// TIA Portal project "Linie_reciclare_paleti_mod" (V16) (continued)
               Length : Int := 1;
               BlockStat : DWord;
               IOLStat : DWord;
               RelRead : Bool := TRUE;
               RelWrite : Bool := TRUE;
            END_STRUCT;
            Parameter_13 : Struct
               V_X1_3_DO2Sub8 : Byte := BYTE#16#00;
               Byte01 : Byte := BYTE#16#00;
               Byte02 : Byte := BYTE#16#00;
               Byte03 : Byte := BYTE#16#00;
               Index : Int := 15000;
               Subindex : Int := 8;
               Length : Int := 1;
               BlockStat : DWord;
               IOLStat : DWord;
               RelRead : Bool := TRUE;
               RelWrite : Bool := TRUE;
            END_STRUCT;
            Parameter_14 : Struct
               V_X1_4_DO1Sub9 : Byte := BYTE#16#00;
               Byte01 : Byte := BYTE#16#00;
               Byte02 : Byte := BYTE#16#00;
               Byte03 : Byte := BYTE#16#00;
               Index : Int := 15000;
               Subindex : Int := 9;
               Length : Int := 1;
               BlockStat : DWord;
               IOLStat : DWord;
               RelRead : Bool := TRUE;
               RelWrite : Bool := TRUE;
            END_STRUCT;
            Parameter_15 : Struct
               V_X1_4_DO2Sub10 : Byte := BYTE#16#00;
               Byte01 : Byte := BYTE#16#00;
               Byte02 : Byte := BYTE#16#00;
               Byte03 : Byte := BYTE#16#00;
               Index : Int := 15000;
               Subindex : Int := 10;
               Length : Int := 1;
               BlockStat : DWord;
               IOLStat : DWord;
               RelRead : Bool := TRUE;
               RelWrite : Bool := TRUE;
            END_STRUCT;
            Parameter_16 : Struct
               V_X1_5_DO1Sub11 : Byte := BYTE#16#00;
               Byte01 : Byte := BYTE#16#00;
               Byte02 : Byte := BYTE#16#00;
               Byte03 : Byte := BYTE#16#00;
               Index : Int := 15000;
               Subindex : Int := 11;
               Length : Int := 1;
               BlockStat : DWord;
               IOLStat : DWord;
               RelRead : Bool := TRUE;
               RelWrite : Bool := TRUE;
            END_STRUCT;
            Parameter_17 : Struct
               V_X1_5_DO2Sub12 : Byte := BYTE#16#00;
               Byte01 : Byte := BYTE#16#00;
               Byte02 : Byte := BYTE#16#00;
               Byte03 : Byte := BYTE#16#00;
               Index : Int := 15000;
               Subindex : Int := 12;
               Length : Int := 1;
               BlockStat : DWord;
               IOLStat : DWord;
               RelRead : Bool := TRUE;
               RelWrite : Bool := TRUE;
            END_STRUCT;
            Parameter_18 : Struct
               V_X1_6_DO1Sub13 : Byte := BYTE#16#80;
               Byte01 : Byte := BYTE#16#00;
               Byte02 : Byte := BYTE#16#00;
               Byte03 : Byte := BYTE#16#00;
               Index : Int := 15000;
               Subindex : Int := 13;
               Length : Int := 1;
               BlockStat : DWord;
               IOLStat : DWord;
               RelRead : Bool := TRUE;
               RelWrite : Bool := TRUE;
            END_STRUCT;
            Parameter_19 : Struct
               V_X1_6_DO2Sub14 : Byte := BYTE#16#80;
               Byte01 : Byte := BYTE#16#00;
               Byte02 : Byte := BYTE#16#00;
               Byte03 : Byte := BYTE#16#00;
               Index : Int := 15000;
               Subindex : Int := 14;
               Length : Int := 1;
               BlockStat : DWord;
               IOLStat : DWord;
               RelRead : Bool := TRUE;
               RelWrite : Bool := TRUE;
            END_STRUCT;
            Parameter_20 : Struct
               V_X1_7_DO1Sub15 : Byte := BYTE#16#80;
               Byte01 : Byte := BYTE#16#00;
               Byte02 : Byte := BYTE#16#00;
               Byte03 : Byte := BYTE#16#00;
               Index : Int := 15000;
               Subindex : Int := 15;
               Length : Int := 1;
               BlockStat : DWord;
               IOLStat : DWord;
               RelRead : Bool := TRUE;
               RelWrite : Bool := TRUE;
            END_STRUCT;
            Parameter_21 : Struct
               V_X1_7_DO2Sub16 : Byte := BYTE#16#80;
               Byte01 : Byte := BYTE#16#00;
               Byte02 : Byte := BYTE#16#00;
               Byte03 : Byte := BYTE#16#00;
               Index : Int := 15000;
               Subindex : Int := 16;
               Length : Int := 1;
               BlockStat : DWord;
               IOLStat : DWord;
               RelRead : Bool := TRUE;
               RelWrite : Bool := TRUE;
            END_STRUCT;
            Parameter_22 : Struct
               V_X1_8_DO1Sub17 : Byte := BYTE#16#80;
               Byte01 : Byte := BYTE#16#00;
               Byte02 : Byte := BYTE#16#00;
               Byte03 : Byte := BYTE#16#00;
               Index : Int := 15000;
               Subindex : Int := 17;
               Length : Int := 1;
               BlockStat : DWord;
               IOLStat : DWord;
               RelRead : Bool := TRUE;
               RelWrite : Bool := TRUE;
            END_STRUCT;
            Parameter_23 : Struct
               V_X1_8_DO2Sub18 : Byte := BYTE#16#80;
               Byte01 : Byte := BYTE#16#00;
               Byte02 : Byte := BYTE#16#00;
               Byte03 : Byte := BYTE#16#00;
               Index : Int := 15000;
               Subindex : Int := 18;
               Length : Int := 1;
               BlockStat : DWord;
               IOLStat : DWord;
               RelRead : Bool := TRUE;
               RelWrite : Bool := TRUE;
            END_STRUCT;
            Parameter_24 : Struct
               V_X1_9_DO1Sub19 : Byte := BYTE#16#80;
               Byte01 : Byte := BYTE#16#00;
               Byte02 : Byte := BYTE#16#00;
               Byte03 : Byte := BYTE#16#00;
               Index : Int := 15000;
               Subindex : Int := 19;
               Length : Int := 1;
               BlockStat : DWord;
               IOLStat : DWord;
               RelRead : Bool := TRUE;
               RelWrite : Bool := TRUE;
            END_STRUCT;
            Parameter_25 : Struct
               V_X1_9_DO2Sub20 : Byte := BYTE#16#80;
               Byte01 : Byte := BYTE#16#00;
               Byte02 : Byte := BYTE#16#00;
               Byte03 : Byte := BYTE#16#00;
               Index : Int := 15000;
               Subindex : Int := 20;
               Length : Int := 1;
               BlockStat : DWord;
               IOLStat : DWord;
               RelRead : Bool := TRUE;
               RelWrite : Bool := TRUE;
            END_STRUCT;
            Parameter_26 : Struct
               V_X1_10_DO1Sub21 : Byte := BYTE#16#80;
               Byte01 : Byte := BYTE#16#00;
               Byte02 : Byte := BYTE#16#00;
               Byte03 : Byte := BYTE#16#00;
               Index : Int := 15000;
               Subindex : Int := 21;
               Length : Int := 1;
               BlockStat : DWord;
               IOLStat : DWord;
               RelRead : Bool := TRUE;
               RelWrite : Bool := TRUE;
            END_STRUCT;
            Parameter_27 : Struct
               V_X1_10_DO2Sub22 : Byte := BYTE#16#80;
               Byte01 : Byte := BYTE#16#00;
               Byte02 : Byte := BYTE#16#00;
               Byte03 : Byte := BYTE#16#00;
               Index : Int := 15000;
               Subindex : Int := 22;
               Length : Int := 1;
               BlockStat : DWord;
               IOLStat : DWord;
               RelRead : Bool := TRUE;
               RelWrite : Bool := TRUE;
            END_STRUCT;
            Parameter_28 : Struct
               V_X1_11_DO1Sub23 : Byte := BYTE#16#80;
               Byte01 : Byte := BYTE#16#00;
               Byte02 : Byte := BYTE#16#00;
               Byte03 : Byte := BYTE#16#00;
               Index : Int := 15000;
               Subindex : Int := 23;
               Length : Int := 1;
               BlockStat : DWord;
               IOLStat : DWord;
               RelRead : Bool := TRUE;
               RelWrite : Bool := TRUE;
            END_STRUCT;
            Parameter_29 : Struct
               V_X1_11_DO2Sub24 : Byte := BYTE#16#80;
               Byte01 : Byte := BYTE#16#00;
               Byte02 : Byte := BYTE#16#00;
               Byte03 : Byte := BYTE#16#00;
               Index : Int := 15000;
               Subindex : Int := 24;
               Length : Int := 1;
               BlockStat : DWord;
               IOLStat : DWord;
               RelRead : Bool := TRUE;
               RelWrite : Bool := TRUE;
            END_STRUCT;
            Parameter_30 : Struct
               V_X1_12_DO1Sub25 : Byte := BYTE#16#80;
               Byte01 : Byte := BYTE#16#00;
               Byte02 : Byte := BYTE#16#00;
               Byte03 : Byte := BYTE#16#00;
               Index : Int := 15000;
               Subindex : Int := 25;
               Length : Int := 1;
               BlockStat : DWord;
               IOLStat : DWord;
               RelRead : Bool := TRUE;
               RelWrite : Bool := TRUE;
            END_STRUCT;
            Parameter_31 : Struct
               V_X1_12_DO2Sub26 : Byte := BYTE#16#80;
               Byte01 : Byte := BYTE#16#00;
               Byte02 : Byte := BYTE#16#00;
               Byte03 : Byte := BYTE#16#00;
               Index : Int := 15000;
               Subindex : Int := 26;
               Length : Int := 1;
               BlockStat : DWord;
               IOLStat : DWord;
               RelRead : Bool := TRUE;
               RelWrite : Bool := TRUE;
            END_STRUCT;
            Parameter_32 : Struct
               V_X1_13_DO1Sub27 : Byte := BYTE#16#80;
               Byte01 : Byte := BYTE#16#00;
               Byte02 : Byte := BYTE#16#00;
               Byte03 : Byte := BYTE#16#00;
               Index : Int := 15000;
               Subindex : Int := 27;
               Length : Int := 1;
               BlockStat : DWord;
               IOLStat : DWord;
               RelRead : Bool := TRUE;
               RelWrite : Bool := TRUE;
            END_STRUCT;
            Parameter_33 : Struct
               V_X1_13_DO2Sub28 : Byte := BYTE#16#80;
               Byte01 : Byte := BYTE#16#00;
               Byte02 : Byte := BYTE#16#00;
               Byte03 : Byte := BYTE#16#00;
               Index : Int := 15000;
               Subindex : Int := 28;
               Length : Int := 1;
               BlockStat : DWord;
               IOLStat : DWord;
               RelRead : Bool := TRUE;
               RelWrite : Bool := TRUE;
            END_STRUCT;
            Parameter_34 : Struct
               V_X1_14_DO1Sub29 : Byte := BYTE#16#80;
               Byte01 : Byte := BYTE#16#00;
               Byte02 : Byte := BYTE#16#00;
               Byte03 : Byte := BYTE#16#00;
               Index : Int := 15000;
               Subindex : Int := 29;
               Length : Int := 1;
               BlockStat : DWord;
               IOLStat : DWord;
               RelRead : Bool := TRUE;
               RelWrite : Bool := TRUE;
            END_STRUCT;
            Parameter_35 : Struct
               V_X1_14_DO2Sub30 : Byte := BYTE#16#80;
               Byte01 : Byte := BYTE#16#00;
               Byte02 : Byte := BYTE#16#00;
               Byte03 : Byte := BYTE#16#00;
               Index : Int := 15000;
               Subindex : Int := 30;
               Length : Int := 1;
               BlockStat : DWord;
               IOLStat : DWord;
               RelRead : Bool := TRUE;
               RelWrite : Bool := TRUE;
            END_STRUCT;
            Parameter_36 : Struct
               V_X1_15_DO1Sub31 : Byte := BYTE#16#80;
               Byte01 : Byte := BYTE#16#00;
               Byte02 : Byte := BYTE#16#00;
               Byte03 : Byte := BYTE#16#00;
               Index : Int := 15000;
               Subindex : Int := 31;
               Length : Int := 1;
               BlockStat : DWord;
               IOLStat : DWord;
               RelRead : Bool := TRUE;
               RelWrite : Bool := TRUE;
            END_STRUCT;
            Parameter_37 : Struct
               V_X1_15_DO2Sub32 : Byte := BYTE#16#80;
               Byte01 : Byte := BYTE#16#00;
               Byte02 : Byte := BYTE#16#00;
               Byte03 : Byte := BYTE#16#00;
               Index : Int := 15000;
               Subindex : Int := 32;
               Length : Int := 1;
               BlockStat : DWord;
               IOLStat : DWord;
               RelRead : Bool := TRUE;
               RelWrite : Bool := TRUE;
            END_STRUCT;
         END_STRUCT;
         Commando : Struct
            Commando_00 : Struct
               Value : Byte := BYTE#16#82;
               Index : Int := 2;
               Subindex : Int := 0;
               Length : Int := 1;
               BlockStat : DWord;
               IOLStat : DWord;
            END_STRUCT;
            Commando_01 : Struct
               Value : Byte := BYTE#16#D0;
               Index : Int := 2;
               Subindex : Int := 0;
               Length : Int := 1;
               BlockStat : DWord;
               IOLStat : DWord;
            END_STRUCT;
            Commando_02 : Struct
               Value : Byte := BYTE#16#D1;
               Index : Int := 2;
               Subindex : Int := 0;
               Length : Int := 1;
               BlockStat : DWord;
               IOLStat : DWord;
            END_STRUCT;
            Commando_03 : Struct
               Value : Byte := BYTE#16#F0;
               Index : Int := 2;
               Subindex : Int := 0;
               Length : Int := 1;
               BlockStat : DWord;
               IOLStat : DWord;
            END_STRUCT;
            Commando_04 : Struct
               Value : Byte := BYTE#16#F1;
               Index : Int := 2;
               Subindex : Int := 0;
               Length : Int := 1;
               BlockStat : DWord;
               IOLStat : DWord;
            END_STRUCT;
            Commando_05 : Struct
               Value : Byte := BYTE#16#F2;
               Index : Int := 2;
               Subindex : Int := 0;
               Length : Int := 1;
               BlockStat : DWord;
               IOLStat : DWord;
            END_STRUCT;
            Commando_06 : Struct
               Value : Byte := BYTE#16#F3;
               Index : Int := 2;
               Subindex : Int := 0;
               Length : Int := 1;
               BlockStat : DWord;
               IOLStat : DWord;
            END_STRUCT;
         END_STRUCT;
      END_STRUCT;
   END_STRUCT;
END_TYPE

TYPE "Bits_Stacker"
VERSION : 0.1
   STRUCT
      Input : Struct
         iEnable : Bool;
         iReset : Bool;
         iAutomatic : Bool;
         iManual : Bool;
         iManualUp : Bool;
         iManualDown : Bool;
         iManualOpenForks : Bool;
         iManualCloseForks : Bool;
         Vertical_sus : Bool;
         Vertical_mijloc : Bool;
         iB10 : Bool;
         Vertical_jos : Bool;
         Furca_extins : Bool;
         Furca_retras : Bool;
         Detectie_palet : Bool;
         Senzor_stiva : Bool;
      END_STRUCT;
      Output : Struct
         Cmd_sus : Bool;
         Cmd_jos : Bool;
         Cmd_extindere : Bool;
         Cmd_retragere : Bool;
         oAlarmUpDown : Bool;
         oAlarmForks : Bool;
         oAlarmPosition : Bool;
         oAlarmFull : Bool;
      END_STRUCT;
   END_STRUCT;
END_TYPE

TYPE "Bits_Drive"
VERSION : 0.1
   STRUCT
      Input : Struct
         iStart : Bool;
         iStop : Bool;
         iProtectie : Bool;
         iContactor : Bool;
         iBrake : Bool;
         iRun : Bool;
         iFault : Bool;
         iReset_Fault : Bool;
         iAckFault : Bool;
      END_STRUCT;
      Output : Struct
         oContactor : Bool;
         oON : Bool;
         oBrake : Bool;
         oFault : Bool;
         oAlarmProtectie : Bool;
         oAlarmContactor : Bool;
         oAlarmBrake : Bool;
         oAckFault : Bool;
      END_STRUCT;
   END_STRUCT;
END_TYPE

TYPE "udt_transit"
VERSION : 0.1
   STRUCT
      trans : Bool;
      alm_tmt : Bool;
      alm_release : Bool;
   END_STRUCT;
END_TYPE

TYPE "Settings_Palletdispenser_PD2"
VERSION : 0.1
   STRUCT
      Configuration : Struct
         Mode : Int := 1;
         Pallettype : Int := 0;
         Double : Bool;
      END_STRUCT;
      MaximumDurationUpDown : DInt := 10000;
      MaximumDurationForks : DInt := 10000;
   END_STRUCT;
END_TYPE

TYPE "udt_step"
VERSION : 0.1
   STRUCT
      wait : Bool;
   END_STRUCT;
END_TYPE

TYPE "MDM"
   STRUCT
      Auto : Bool;
      Manual : Bool;
      "Step" : Bool;
      Start : Bool;
      Stop : Bool;
   END_STRUCT;
END_TYPE

TYPE "Handshakes_PalletDispenser_PD2"
VERSION : 0.1
   STRUCT
      Command : Struct
         Deliver : Bool;
         PickUpStack : Bool;
         WaitPosition : Bool;
         Receive : Bool;
         Pallettype : Int;
      END_STRUCT;
      Status : Struct
         Blocked : Bool;
         PalletPresent : Bool;
         BasicPosition : Bool;
         WaitPosition : Bool;
         Busy : Bool;
         Pallettype : Int;
         "Step" : Int;
      END_STRUCT;
   END_STRUCT;
END_TYPE

DATA_BLOCK "DB2_WORK_BITS"   // DB2
{ S7_Optimized_Access := 'TRUE' }
VERSION : 0.1
   VAR
      Settings_DeStacker : "Settings_Palletdispenser_PD2";
      Handshakes_DeStacker : "Handshakes_PalletDispenser_PD2";
      Settings_Destacker_Finished : Bool;
      Stacker_New_Handler : "Bits_Stacker";
      SQ_Outfeed_Stack_SN : Bool;
      Pallet_fed : Bool;
      Start_Destacker_Cycle : Bool;
      Enable_Destacker : Bool;
      Destacker_Busy_Timer : Time;
      SQ_Pallet_Length_Stacker_New : Bool;
      Pallet_Length_Stacker_New : Int;
      SQ_Pallet_Length_Stacker : Bool;
      Pallet_Length_Stacker : Int;
      SQ_SN_Length : Array[0..2] of Bool;
      SQ_S_Length : Array[0..2] of Bool;
      Length : Struct
         Length_1 : Array[0..2] of Int;
         Length_2 : Array[0..2] of Int;
         Length_3 : Array[0..2] of Int;
      END_STRUCT;
      DS_Stop_Drive : Bool;
      S_Stop_Drive : Bool;
      Settings_Stacker_Finished : Bool;
      Settings_Stacker : "Settings_Palletdispenser_PD2";
      Settings_Stacker_New : "Settings_Palletdispenser_PD2";
      Stacker_Handler : "Bits_Stacker";
      Handshakes_Stacker : "Handshakes_PalletDispenser_PD2";
      Handshakes_Stacker_New : "Handshakes_PalletDispenser_PD2";
      Enable_Stacker : Bool;
      Sart_Stacker_Cycle : Bool;
      SQ_Outfeed_Stack_S : Bool;
      Stack_fed : Bool;
      Stacker_Busy_Timer : Time;
      Stacker_New_Drive_Handler : "Bits_Drive";
      Stacker_Drive_Handler : "Bits_Drive";
      CD_Drive_Handler : "Bits_Drive";
      Operating_Modes : Struct
         Automatic : Bool := true;
         Maintenance : Bool;
      END_STRUCT;
      DS_Machine_Checked : Bool;
      SQs_Loading_Stack : Struct
         SQ_Stack_Present : Bool;
         SQ_Stack_Height : Bool;
         SQ_Left_Align : Bool;
         SQ_Right_Align_1 : Bool;
         SQ_Right_Align_2 : Bool;
      END_STRUCT;
      LStack_OK : Bool;
      Stack_On_Conveyor : Bool;
      SoftStart_Stacker_Nou : Struct
         YV1 : Bool;
         YV2 : Bool;
         Sensor1 : Bool;
         Sensor2 : Bool;
      END_STRUCT;
      SoftStart_Stacker : Struct
         YV1 : Bool;
         YV2 : Bool;
         Sensor1 : Bool;
         Sensor2 : Bool;
      END_STRUCT;
      SoftStart_Zone2_A : Struct
         YV1 : Bool;
         YV2 : Bool;
         Sensor1 : Bool;
         Sensor2 : Bool;
      END_STRUCT;
      SoftStart_Zone2_B : Struct
         YV1 : Bool;
         YV2 : Bool;
         Sensor1 : Bool;
         Sensor2 : Bool;
      END_STRUCT;
      Motor_Transport_S : Struct
         ON : Bool;
         RUN : Bool;
         Protectie : Bool;
      END_STRUCT;
      Motor_Transport_SN : Struct
         ON : Bool;
         RUN : Bool;
         Protectie : Bool;
      END_STRUCT;
      Motor_Centror_S : Struct
         ON : Bool;
         RUN : Bool;
         Protectie : Bool;
      END_STRUCT;
      Motor_Centror_SN : Struct
         ON : Bool;
         RUN : Bool;
         Protectie : Bool;
      END_STRUCT;
      Transport_Conveyor_SQs : Struct
         SQ_Repaired_Pallet : Array[0..1] of Bool;
         SQ_Conveyor_End : Bool;
      END_STRUCT;
      SQ_Centror_S : Bool;
      SQ_Centror_SN : Bool;
      Centror_S : Struct
         YV_centror_centr : Bool;
         YV_centror_eliber : Bool;
         Sensor_eliber : Bool;
         Sensor_centr : Bool;
         Centered : Bool;
      END_STRUCT;
      Centror_SN : Struct
         YV_centror_centr : Bool;
         YV_centror_eliber : Bool;
         Sensor_eliber : Bool;
         Sensor_centr : Bool;
         Centered : Bool;
      END_STRUCT;
      Stack_Output_Drive_Handler : "Bits_Drive";
      Stack_New_Output_Drive_Handler : "Bits_Drive";
      Stacker_Full : Bool;
      AG : Struct
         Air : Bool;
         Ilum : Bool;
         Fixed_Saw : Bool;
         HMI : Bool;
         MDP_S : Bool;
         MDP_D : Bool;
         "PR_S+D" : Bool;
         PR_M : Bool;
         TELE : Bool;
      END_STRUCT;
      AG_Lamp : Struct
         Red : Bool;
         Yellow : Bool;
         Green : Bool;
      END_STRUCT;
      Previous_Length : Int;
      Same_Length : Bool;
      BDS : Struct
         Red : Bool;
         Yellow : Bool;
         Green : Bool;
      END_STRUCT;
      BS : Struct
         Red : Bool;
         Yellow : Bool;
         Green : Bool;
      END_STRUCT;
      Consumption_Pulse : Bool;
      Start : Bool;
      Conveyor_Speed_SN : Int := 398;
      Stops : Struct
         DS : Bool;
         S : Bool;
      END_STRUCT;
      DS_Waiting : Bool;
      RS_DS : Bool;   // Comanda Cilindru JOS
      Conveyor_Speed_S : Int := 1200;
      Switch_output : Bool;
      LED : Bool;
      Reset_S : Struct
         Up : Bool;
         Down : Bool;
         InStack : Bool;
         OutStack : Bool;
      END_STRUCT;
      Reset_DS : Struct
         Up : Bool;
         Down : Bool;
         InStack : Bool;
         OutStack : Bool;
      END_STRUCT;
      Reset_LED_Count : Bool;
      Start_ON : Bool;
      DS_Step3_OK : Bool;
      Reset_Clock_SN : Bool;
      Reset_Counter_SN : Bool;
      Reset_Clock_S : Bool;
      Reset_Counter_S : Bool;
      Synth_Alarms : Bool;
      Ton : Array[0..30] of TON_TIME;
      Select_MDM : Int;
      MDM : Array[0..1] of "MDM";
   END_VAR
BEGIN
   Length.Length_1[0] := 1000;
   Length.Length_1[1] := 1100;
   Length.Length_1[2] := 1350;
   Length.Length_2[0] := 1600;
   Length.Length_2[1] := 1500;
   Length.Length_2[2] := 1700;
   Length.Length_3[0] := 2000;
   Length.Length_3[1] := 1900;
   Length.Length_3[2] := 2500;
   Settings_Stacker.Configuration.Mode := 2;
   Settings_Stacker_New.Configuration.Mode := 2;
   // MDM[0] : Line A
   // MDM[1] : Line B
END_DATA_BLOCK

DATA_BLOCK "DB3_FAULTS"   // DB3
{ S7_Optimized_Access := 'FALSE' }
VERSION : 0.1
   VAR
      Safety_Synth_SN : Bool;
      Safety_Synth_Zone2 : Bool;
      Safety_Synth_S : Bool;
      Alarm_Stacker_New : Word;
      Fault_Pallet_Length_Stacker_New : Bool;
      Fault_Pallet_Length_Stacker : Bool;
      Alarm_Stacker : Word;
      Alarm_Centror : Word;
      Alarm_CD1 : Word;
      Alarm_CD2 : Word;
      Alarm_CS1 : Word;
      Alarm_CS2 : Word;
      Alarm_CS3 : Word;
      Alarm_CS4 : Word;
      Alarm_Safety_SN : Word;
      Alarm_Safety_Z2 : Word;
      Alarm_Safety_S : Word;
      Alarm_General_S : Word;
      Alarm_General_SN : Word;
   END_VAR
BEGIN
END_DATA_BLOCK

DATA_BLOCK "FB_Pallet_Length_DB_Stacker"   // DB6
{ S7_Optimized_Access := 'TRUE' }
VERSION : 0.1
// stored: InstanceOfName FB_Pallet_Length
"FB_Pallet_Length"
BEGIN
END_DATA_BLOCK

DATA_BLOCK "DB_DRIVE_DESTACKER"   // DB10
{ S7_Optimized_Access := 'TRUE' }
VERSION : 0.1
// stored: InstanceOfName FB1_DRIVE
"FB1_DRIVE"
BEGIN
END_DATA_BLOCK

DATA_BLOCK "DB_DRIVE_CD"   // DB12
{ S7_Optimized_Access := 'TRUE' }
VERSION : 0.1
// stored: InstanceOfName FB1_DRIVE
"FB1_DRIVE"
BEGIN
END_DATA_BLOCK

DATA_BLOCK "FB_DS_Check_Machine_DB"   // DB14
{ S7_Optimized_Access := 'TRUE' }
VERSION : 0.1
// stored: InstanceOfName FB_DS_Check_Machine
"FB_DS_Check_Machine"
BEGIN
END_DATA_BLOCK

DATA_BLOCK "DB_DRIVE_STACKER"   // DB17
{ S7_Optimized_Access := 'TRUE' }
VERSION : 0.1
// stored: InstanceOfName FB1_DRIVE
"FB1_DRIVE"
BEGIN
END_DATA_BLOCK

DATA_BLOCK "DB_DRIVE_STACK_OUTPUT"   // DB18
{ S7_Optimized_Access := 'TRUE' }
VERSION : 0.1
// stored: InstanceOfName FB1_DRIVE
"FB1_DRIVE"
BEGIN
END_DATA_BLOCK

DATA_BLOCK "FB_EnergyCounter_DB"   // DB19
{ S7_Optimized_Access := 'TRUE' }
VERSION : 0.1
// stored: InstanceOfName FB_EnergyCounter
"FB_EnergyCounter"
BEGIN
END_DATA_BLOCK

DATA_BLOCK "DB20_DATA_HMI"   // DB20
{ S7_Optimized_Access := 'TRUE' }
VERSION : 0.1
   VAR
      Reset_Faults : Bool;
      Destacker_Manual : Struct
         Up : Bool;
         Down : Bool;
         Extend : Bool;
         Retract : Bool;
      END_STRUCT;
      Stacker_Manual : Struct
         Up : Bool;
         Down : Bool;
         Extend : Bool;
         Retract : Bool;
      END_STRUCT;
      Run : Bool;
      Maintenance : Bool;
      Conveyors_Manual : Struct
         CD1 : Bool;
         CD2 : Bool;
         T : Bool;
         C : Bool;
         CS1 : Bool;
         CS2 : Bool;
      END_STRUCT;
      Step_Destacker : Int;
      Step_Stacker : Int;
   END_VAR
BEGIN
END_DATA_BLOCK

DATA_BLOCK "FB_AlarmCounter_DB"   // DB22
{ S7_Optimized_Access := 'TRUE' }
VERSION : 0.1
// stored: InstanceOfName FB_AlarmCounter
"FB_AlarmCounter"
BEGIN
END_DATA_BLOCK

DATA_BLOCK "FB_IntervalTrigger_DB"   // DB23
{ S7_Optimized_Access := 'TRUE' }
VERSION : 0.1
// stored: InstanceOfName FB_IntervalTrigger
"FB_IntervalTrigger"
BEGIN
END_DATA_BLOCK

DATA_BLOCK "DB29_SECU_OUT"   // DB29
{ S7_Optimized_Access := 'TRUE' }
VERSION : 0.1
   VAR
      Reset_DS_Relay : Bool;
      Reset_DS_Barrier : Bool;
      Reset_Z2_Relay : Bool;
      Reset_S_Relay : Bool;
      Reset_S_Barrier_1 : Bool;
      Reset_S_Barrier_2 : Bool;
   END_VAR
BEGIN
END_DATA_BLOCK

DATA_BLOCK "O"   // DB30
{ S7_Optimized_Access := 'TRUE' }
VERSION : 0.1
// stored: InstanceOfName FB_Outputs
"FB_Outputs"
BEGIN
END_DATA_BLOCK

DATA_BLOCK "FB_ProductionStatistics_DB"   // DB31
{ S7_Optimized_Access := 'TRUE' }
VERSION : 0.1
// stored: InstanceOfName FB_ProductionStatistics
"FB_ProductionStatistics"
BEGIN
END_DATA_BLOCK

DATA_BLOCK "DB_Init_S"   // DB35
{ S7_Optimized_Access := 'TRUE' }
VERSION : 0.1
// stored: InstanceOfName FB_Init_S
"FB_Init_S"
BEGIN
END_DATA_BLOCK

DATA_BLOCK "DB_Centrare"   // DB36
{ S7_Optimized_Access := 'TRUE' }
VERSION : 0.1
// stored: InstanceOfName FB_Centrare
"FB_Centrare"
BEGIN
END_DATA_BLOCK

DATA_BLOCK "DB_MDM_S"   // DB37
{ S7_Optimized_Access := 'TRUE' }
VERSION : 0.1
// stored: InstanceOfName FB_MDM
"FB_MDM"
BEGIN
END_DATA_BLOCK

DATA_BLOCK "st"   // DB39
{ S7_Optimized_Access := 'TRUE' }
VERSION : 0.1
// stored: InstanceOfName FB_MDM
"FB_MDM"
BEGIN
END_DATA_BLOCK

DATA_BLOCK "s"   // DB40
{ S7_Optimized_Access := 'TRUE' }
VERSION : 0.1
// stored: InstanceOfName StaCall
"StaCall"
BEGIN
   nAc := 2;
END_DATA_BLOCK

DATA_BLOCK "ds"   // DB41
{ S7_Optimized_Access := 'TRUE' }
VERSION : 0.1
// stored: InstanceOfName StaCall
"StaCall"
BEGIN
END_DATA_BLOCK

DATA_BLOCK "x"   // DB43
{ S7_Optimized_Access := 'TRUE' }
VERSION : 0.1
   VAR
      "b" : Array[0..31] of Bool;
      f : Array[0..31] of Bool;
      bs : Array[0..10] of SInt;
      bt : Array[0..10] of SInt;
      set_Bk_all : Bool;
      rset_Bk_all : Bool;
      stp_Bk_s : Bool;
      stp_Bk_En : Bool;
      stp_Bk_t : Bool;
      stp_Bk_c : Bool;
      dlyt : Array[0..10] of Bool;
      wd : Array[0..10] of Int;
      dlyc : Array[0..10] of SInt;
      bkS_Adm : Array[0..9] of Bool;
      bkS_Eva : Array[0..9] of Bool;
      bkC_Av : Array[0..9] of Bool;
      bkC_Ret : Array[0..9] of Bool;
      evac : Array[0..7] of Bool;
      bb : Array[0..31] of Bool;
   END_VAR
BEGIN
END_DATA_BLOCK

DATA_BLOCK "alm"   // DB44
{ S7_Optimized_Access := 'FALSE' }
VERSION : 0.1
   VAR
      alms : Array[0..9] of SInt;
      almt : Array[0..9] of SInt;
      almc : Array[0..9] of SInt;
      alms_dis : Array[0..9] of SInt;
      almt_dis : Array[0..9] of SInt;
      almc_dis : Array[0..9] of SInt;
      alms_m : Array[0..9] of SInt;
      almt_m : Array[0..9] of SInt;
      almc_m : Array[0..9] of SInt;
      almsf : Array[0..4] of SInt;
      almr : Array[0..4] of SInt;
   END_VAR
BEGIN
   almt_dis[1] := 3;
END_DATA_BLOCK

DATA_BLOCK "Gen"   // DB45
{ S7_Optimized_Access := 'TRUE' }
VERSION : 0.1
   VAR RETAIN
      optConvIn : Bool;   // 0-Conv In liber 1-Conv In comandat de lant
   END_VAR
   VAR
      tct : UInt;
      tctv : UInt;
      tctf : UInt;
      tm1s : IEC_TIMER;
      ModNoSafe : Bool;
      ModEnergie : Bool;
      "Mod Man" : Bool;
      ModWait : Bool;
      ModInit : Bool;
      ModAuto : Bool;
      ModCycle : Bool;
      ModPas : Bool;
      AlarmStop : Bool;
      AlarmRun : Bool;
      ButResetAlarm : Bool;
      ButResetSafe : Bool;
      ButInit : Bool;
      ButStartCycle : Bool;
      ButStopCycle : Bool;
      ButStopCycleEnd : Bool;
      ButAuto : Bool;
      ButStep : Bool;
      StepMod : UInt;
      StepModImg : UInt;
      Safe : Bool;
      Init_OK : Bool;
      SafeConv : Bool;
      PowerConv : Bool;
      Energy : Bool;
   END_VAR
   VAR RETAIN
      optAckOp : Bool;
   END_VAR
   VAR
      S_AlarmAny : Bool;
      SN_AlarmAny : Bool;
      Ton : Array[0..20] of IEC_TIMER;
   END_VAR
BEGIN
END_DATA_BLOCK

DATA_BLOCK "HMI"   // DB46
{ S7_Optimized_Access := 'FALSE' }
VERSION : 0.1
   VAR
      popupEn : Array[0..9] of Bool;
      popupMsj : Array[0..9] of USInt;
      spare : Array[0..4] of USInt;
      pg : Array[0..7] of USInt;
      pg_cfg : Array[0..7] of USInt;
      statie_sel : Int;
      tranzit_sel : Int;
      cil_sel : Int;
      tip_sel : Int;
      instance_sel : Int;
      numSt : USInt;
      numSt_s : USInt;
      numCyl : USInt;
      numSens : USInt;
      pgCfg : USInt;
      pgCfgV : USInt;
      ButOpVis : USInt;
      ButOp : Array[0..7] of Bool;
      tip_sel_v : Int;
      instance_sel_v : Int;
      chg_prio : Bool;
      ButOpMem : USInt;
      ButOpW : USInt;
      ButOpHMI : USInt;
      msop_vizi : USInt;
      msop_NoAlm : Bool;
      hmi_stat_arrow : Array[0..10] of USInt;
      CfOp : Array[0..31] of Bool;
   END_VAR
BEGIN
END_DATA_BLOCK

DATA_BLOCK "Cylinder_la_in"   // DB47
{ S7_Optimized_Access := 'TRUE' }
VERSION : 0.1
// stored: InstanceOfName Cylinder
"Cylinder"
BEGIN
END_DATA_BLOCK

DATA_BLOCK "Cylinder_la_out"   // DB48
{ S7_Optimized_Access := 'TRUE' }
VERSION : 0.1
// stored: InstanceOfName Cylinder
"Cylinder"
BEGIN
END_DATA_BLOCK

DATA_BLOCK "Cylinder_GripV_M"   // DB49
{ S7_Optimized_Access := 'TRUE' }
VERSION : 0.1
// stored: InstanceOfName Cylinder
"Cylinder"
BEGIN
END_DATA_BLOCK

DATA_BLOCK "DB50_PALLET_LENGTH"   // DB50
{ S7_Optimized_Access := 'TRUE' }
VERSION : 0.1
BEGIN
END_DATA_BLOCK

DATA_BLOCK "Cylinder_GripH_M"   // DB51
{ S7_Optimized_Access := 'TRUE' }
VERSION : 0.1
// stored: InstanceOfName Cylinder
"Cylinder"
BEGIN
END_DATA_BLOCK

DATA_BLOCK "Cylinder_GripV_E"   // DB52
{ S7_Optimized_Access := 'TRUE' }
VERSION : 0.1
// stored: InstanceOfName Cylinder
"Cylinder"
BEGIN
END_DATA_BLOCK

DATA_BLOCK "Cylinder_GripH_E"   // DB53
{ S7_Optimized_Access := 'TRUE' }
VERSION : 0.1
// stored: InstanceOfName Cylinder
"Cylinder"
BEGIN
END_DATA_BLOCK

DATA_BLOCK "sim_DB"   // DB54
{ S7_Optimized_Access := 'TRUE' }
VERSION : 0.1
// stored: InstanceOfName sim
"sim"
BEGIN
END_DATA_BLOCK

DATA_BLOCK "FB_GEN_DB"   // DB58
{ S7_Optimized_Access := 'TRUE' }
VERSION : 0.1
// stored: InstanceOfName FB_GEN
"FB_GEN"
BEGIN
END_DATA_BLOCK

DATA_BLOCK "t"   // DB59
{ S7_Optimized_Access := 'TRUE' }
VERSION : 0.1
   VAR
      tmr : Array[0..20] of IEC_TIMER;
   END_VAR
BEGIN
END_DATA_BLOCK

DATA_BLOCK "DB_Init_SN"   // DB60
{ S7_Optimized_Access := 'TRUE' }
VERSION : 0.1
// stored: InstanceOfName FB_Init_SN
"FB_Init_SN"
BEGIN
END_DATA_BLOCK

DATA_BLOCK "DB120_GRAFCETS"   // DB120
{ S7_Optimized_Access := 'TRUE' }
VERSION : 0.1
   VAR
      G7_STOP_SN : Int;
      G7_STOP_S : Int;
      G7_RUN_SN : Int;
      G7_RUN_S : Int;
      S_Last_Step : Int;
      SN_Last_Step : Int;
      G7_STOP_Z2 : Int;
      G7_RUN_Z2 : Int;
      G7_Stack : Int;
      G7_Stack_New : Int;
   END_VAR
BEGIN
END_DATA_BLOCK

DATA_BLOCK "DB121_GRAFCETS_COPY"   // DB121
{ S7_Optimized_Access := 'FALSE' }
VERSION : 0.1
   VAR
      G7_STOP_DS : Array[0..31] of Bool;
      G7_STOP_S : Array[0..31] of Bool;
      G7_RUN_DS : Array[0..31] of Bool;
      G7_RUN_S : Array[0..31] of Bool;
   END_VAR
BEGIN
END_DATA_BLOCK

DATA_BLOCK "DB200_SAFETY"   // DB200
{ S7_Optimized_Access := 'FALSE' }
VERSION : 0.1
   VAR
      Main_Door : Bool;
      "E-STOP_SN" : Bool;
      Rearm_SN_Barrier : Bool;
      Rearm_SN_Relay : Bool;
      "E-STOP_Zone2_MBS" : Bool;
      "E-STOP_Zone2_MBD" : Bool;
      "E-STOP_Zone2_B" : Bool;
      "E-STOP_S" : Bool;
      Mutting_Barrier_SN : Bool;
      Safety_Barrier_2_SN_ARMED : Bool;
      Door_S : Bool;
      Mutting_Barrier_S : Bool;
      Rearm_S : Bool;
      Rearm_Zone2A : Bool;
      Rearm_Zone2B : Bool;
      Zone2_Synth : Bool;
      "E-Stop_LineB" : Bool;
      Door_SN : Bool;
      "E-Stop_LineA" : Bool;
      Zone2B_Relay : Bool;
   END_VAR
BEGIN
END_DATA_BLOCK

DATA_BLOCK "DB_PalletDispenser_PD2_Stacking_DB"   // DB301
{ S7_Optimized_Access := 'TRUE' }
VERSION : 0.1
// stored: InstanceOfName FB_PalletDispenser_PD2_Stacking
"FB_PalletDispenser_PD2_Stacking"
BEGIN
END_DATA_BLOCK

// folder: Stacker_New

DATA_BLOCK "DB_Centrare_SN"   // DB4
{ S7_Optimized_Access := 'TRUE' }
VERSION : 0.1
// stored: InstanceOfName FB_Centrare
"FB_Centrare"
BEGIN
END_DATA_BLOCK

DATA_BLOCK "FB_Pallet_Length_DB_Stacker_New"   // DB5
{ S7_Optimized_Access := 'TRUE' }
VERSION : 0.1
// stored: InstanceOfName FB_Pallet_Length
"FB_Pallet_Length"
BEGIN
END_DATA_BLOCK

DATA_BLOCK "x_SN"   // DB61
{ S7_Optimized_Access := 'TRUE' }
VERSION : 0.1
   VAR
      "b" : Array[0..31] of Bool;
      f : Array[0..31] of Bool;
      bs : Array[0..10] of SInt;
      bt : Array[0..10] of SInt;
      set_Bk_all : Bool;
      rset_Bk_all : Bool;
      stp_Bk_s : Bool;
      stp_Bk_En : Bool;
      stp_Bk_t : Bool;
      stp_Bk_c : Bool;
      dlyt : Array[0..10] of Bool;
      wd : Array[0..10] of Int;
      dlyc : Array[0..10] of SInt;
      bkS_Adm : Array[0..9] of Bool;
      bkS_Eva : Array[0..9] of Bool;
      bkC_Av : Array[0..9] of Bool;
      bkC_Ret : Array[0..9] of Bool;
      evac : Array[0..7] of Bool;
      bb : Array[0..31] of Bool;
   END_VAR
BEGIN
END_DATA_BLOCK

DATA_BLOCK "sn"   // DB62
{ S7_Optimized_Access := 'TRUE' }
VERSION : 0.1
// stored: InstanceOfName StaCall_SN
"StaCall_SN"
BEGIN
END_DATA_BLOCK

DATA_BLOCK "DB_MDM_SN"   // DB63
{ S7_Optimized_Access := 'TRUE' }
VERSION : 0.1
// stored: InstanceOfName FB_MDM
"FB_MDM"
BEGIN
END_DATA_BLOCK

DATA_BLOCK "HMI_SN"   // DB64
{ S7_Optimized_Access := 'FALSE' }
VERSION : 0.1
   VAR
      popupEn : Array[0..9] of Bool;
      popupMsj : Array[0..9] of USInt;
      spare : Array[0..4] of USInt;
      pg : Array[0..7] of USInt;
      pg_cfg : Array[0..7] of USInt;
      statie_sel : Int;
      tranzit_sel : Int;
      cil_sel : Int;
      tip_sel : Int;
      instance_sel : Int;
      numSt : USInt;
      numSt_s : USInt;
      numCyl : USInt;
      numSens : USInt;
      pgCfg : USInt;
      pgCfgV : USInt;
      ButOpVis : USInt;
      ButOp : Array[0..7] of Bool;
      tip_sel_v : Int;
      instance_sel_v : Int;
      chg_prio : Bool;
      ButOpMem : USInt;
      ButOpW : USInt;
      ButOpHMI : USInt;
      msop_vizi : USInt;
      msop_NoAlm : Bool;
      hmi_stat_arrow : Array[0..10] of USInt;
      CfOp : Array[0..31] of Bool;
   END_VAR
BEGIN
END_DATA_BLOCK

DATA_BLOCK "DB_PalletDispenser_PD2_Stacking_New_DB"   // DB302
{ S7_Optimized_Access := 'TRUE' }
VERSION : 0.1
// stored: InstanceOfName FB_PalletDispenser_PD2_Stacking
"FB_PalletDispenser_PD2_Stacking"
BEGIN
END_DATA_BLOCK

// folder: System blocks/Program resources

DATA_BLOCK "Counter_Reset_Pallet_SN"   // DB1
{ S7_Optimized_Access := 'TRUE' }
AUTHOR : Simatic
FAMILY : IEC
NAME : CNTR
VERSION : 1.0
// stored: InstanceOfName IEC_COUNTER
"IEC_COUNTER"
BEGIN
END_DATA_BLOCK

DATA_BLOCK "Timer_Brake_Release"   // DB9
{ S7_Optimized_Access := 'TRUE' }
AUTHOR : Simatic
FAMILY : IEC
NAME : IEC_TMR
VERSION : 1.0
// stored: InstanceOfName IEC_TIMER
"IEC_TIMER"
BEGIN
END_DATA_BLOCK

DATA_BLOCK "Timer_Contactor_Drive"   // DB11
{ S7_Optimized_Access := 'TRUE' }
AUTHOR : Simatic
FAMILY : IEC
NAME : IEC_TMR
VERSION : 1.0
// stored: InstanceOfName IEC_TIMER
"IEC_TIMER"
BEGIN
END_DATA_BLOCK

DATA_BLOCK "Timer_Drive_Blocked"   // DB13
{ S7_Optimized_Access := 'TRUE' }
AUTHOR : Simatic
FAMILY : IEC
NAME : IEC_TMR
VERSION : 1.0
// stored: InstanceOfName IEC_TIMER
"IEC_TIMER"
BEGIN
END_DATA_BLOCK

DATA_BLOCK "tmrCkFull"   // DB15
{ S7_Optimized_Access := 'TRUE' }
AUTHOR : Simatic
FAMILY : IEC
NAME : IEC_TMR
VERSION : 1.0
// stored: InstanceOfName IEC_TIMER
"IEC_TIMER"
BEGIN
END_DATA_BLOCK

DATA_BLOCK "IEC_Timer_Start_Motor_Transport"   // DB16
{ S7_Optimized_Access := 'TRUE' }
AUTHOR : Simatic
FAMILY : IEC
NAME : IEC_TMR
VERSION : 1.0
// stored: InstanceOfName IEC_TIMER
"IEC_TIMER"
BEGIN
END_DATA_BLOCK

DATA_BLOCK "Counter_Reset_Pallet_S"   // DB25
{ S7_Optimized_Access := 'TRUE' }
AUTHOR : Simatic
FAMILY : IEC
NAME : CNTR
VERSION : 1.0
// stored: InstanceOfName IEC_COUNTER
"IEC_COUNTER"
BEGIN
END_DATA_BLOCK

DATA_BLOCK "Timer_Start_Centror"   // DB26
{ S7_Optimized_Access := 'TRUE' }
AUTHOR : Simatic
FAMILY : IEC
NAME : IEC_TMR
VERSION : 1.0
// stored: InstanceOfName IEC_TIMER
"IEC_TIMER"
BEGIN
END_DATA_BLOCK

DATA_BLOCK "Timer_Stop_Count_Length"   // DB28
{ S7_Optimized_Access := 'TRUE' }
AUTHOR : Simatic
FAMILY : IEC
NAME : IEC_TMR
VERSION : 1.0
// stored: InstanceOfName IEC_TIMER
"IEC_TIMER"
BEGIN
END_DATA_BLOCK

DATA_BLOCK "tim[5]"   // DB57
{ S7_Optimized_Access := 'TRUE' }
AUTHOR : Simatic
FAMILY : IEC
NAME : IEC_TMR
VERSION : 1.0
// stored: InstanceOfName IEC_TIMER
"IEC_TIMER"
BEGIN
END_DATA_BLOCK

// folder: log

DATA_BLOCK "ms"   // DB27
{ S7_Optimized_Access := 'TRUE' }
VERSION : 0.1
   VAR RETAIN
      tv : Array[0..99] of UInt;
      tvv : Array[0..99] of UInt;
   END_VAR
   VAR
      trig : Int := 0;
   END_VAR
   VAR RETAIN
      i : Int := 1076;
   END_VAR
   VAR
      ivv : Int := 0;
      v : UDInt := 13011;
      cyc : UDInt := 1;
      tim : UDInt := 735;
      vv : UDInt := 49013011;
      spare : Array[0..30] of UInt;
      p1min : Bool := FALSE;
      p100ms : Bool := FALSE;
      c : Int := 0;
      cc : Int := 0;
      ccc : USInt := 0;
      cach : Bool := FALSE;
      cfis : UInt := 0;
      ctrig : UInt := 0;
      tach : IEC_TIMER;
      T_100ms : IEC_TIMER;
      en : Bool := FALSE;
      ir : Int;
      rv : Array[0..10] of UInt;
      rvv : Array[0..10] of UInt;
      vr : UDInt;
      rtr : UDInt;
   END_VAR
BEGIN
   tv[0] := 0;
   tv[1] := 0;
   tv[2] := 1;
   tv[3] := 128;
   tv[4] := 0;
   tv[5] := 0;
   tv[6] := 0;
   tv[7] := 0;
   tv[8] := 0;
   tv[9] := 0;
   tv[10] := 1;
   tv[11] := 13;
   tv[12] := 23;
   tv[13] := 11;
   tv[14] := 0;
   tv[15] := 0;
   tv[16] := 0;
   tv[17] := 0;
   tv[18] := 0;
   tv[19] := 0;
   tv[20] := 0;
   tv[21] := 0;
   tv[22] := 0;
   tv[23] := 0;
   tv[24] := 0;
   tv[25] := 0;
   tv[26] := 0;
   tv[27] := 0;
   tv[28] := 0;
   tv[29] := 0;
   tv[30] := 0;
   tv[31] := 0;
   tv[32] := 0;
   tv[33] := 0;
   tv[34] := 0;
   tv[35] := 0;
   tv[36] := 0;
   tv[37] := 0;
   tv[38] := 0;
   tv[39] := 0;
   tv[40] := 0;
   tv[41] := 0;
   tv[42] := 0;
   tv[43] := 0;
   tv[44] := 0;
   tv[45] := 0;
   tv[46] := 0;
   tv[47] := 0;
   tv[48] := 0;
   tv[49] := 0;
   tv[50] := 0;
   tv[51] := 0;
   tv[52] := 0;
   tv[53] := 0;
   tv[54] := 0;
   tv[55] := 0;
   tv[56] := 0;
   tv[57] := 0;
   tv[58] := 0;
   tv[59] := 0;
   tv[60] := 0;
   tv[61] := 0;
   tv[62] := 0;
   tv[63] := 0;
   tv[64] := 0;
   tv[65] := 0;
   tv[66] := 0;
   tv[67] := 0;
   tv[68] := 0;
   tv[69] := 0;
   tv[70] := 0;
   tv[71] := 0;
   tv[72] := 0;
   tv[73] := 0;
   tv[74] := 0;
   tv[75] := 0;
   tv[76] := 0;
   tv[77] := 0;
   tv[78] := 0;
   tv[79] := 0;
   tv[80] := 0;
   tv[81] := 0;
   tv[82] := 0;
   tv[83] := 0;
   tv[84] := 0;
   tv[85] := 0;
   tv[86] := 0;
   tv[87] := 0;
   tv[88] := 0;
   tv[89] := 0;
   tv[90] := 0;
   tv[91] := 0;
   tv[92] := 0;
   tv[93] := 0;
   tv[94] := 0;
   tv[95] := 0;
   tv[96] := 0;
   tv[97] := 0;
   tv[98] := 0;
   tv[99] := 0;
   tvv[0] := 0;
   tvv[1] := 0;
   tvv[2] := 1;
   tvv[3] := 128;
   tvv[4] := 0;
   tvv[5] := 0;
   tvv[6] := 0;
   tvv[7] := 0;
   tvv[8] := 0;
   tvv[9] := 0;
   tvv[10] := 1;
   tvv[11] := 13;
   tvv[12] := 23;
   tvv[13] := 11;
   tvv[14] := 0;
   tvv[15] := 0;
   tvv[16] := 0;
   tvv[17] := 0;
   tvv[18] := 0;
   tvv[19] := 0;
   tvv[20] := 0;
   tvv[21] := 0;
   tvv[22] := 0;
   tvv[23] := 0;
   tvv[24] := 0;
   tvv[25] := 0;
   tvv[26] := 0;
   tvv[27] := 0;
   tvv[28] := 0;
   tvv[29] := 0;
   tvv[30] := 0;
   tvv[31] := 0;
   tvv[32] := 0;
   tvv[33] := 0;
   tvv[34] := 0;
   tvv[35] := 0;
   tvv[36] := 0;
   tvv[37] := 0;
   tvv[38] := 0;
   tvv[39] := 0;
   tvv[40] := 0;
   tvv[41] := 0;
   tvv[42] := 0;
   tvv[43] := 0;
   tvv[44] := 0;
   tvv[45] := 0;
   tvv[46] := 0;
   tvv[47] := 0;
   tvv[48] := 0;
   tvv[49] := 0;
   tvv[50] := 0;
   tvv[51] := 0;
   tvv[52] := 0;
   tvv[53] := 0;
   tvv[54] := 0;
   tvv[55] := 0;
   tvv[56] := 0;
   tvv[57] := 0;
   tvv[58] := 0;
   tvv[59] := 0;
   tvv[60] := 0;
   tvv[61] := 0;
   tvv[62] := 0;
   tvv[63] := 0;
   tvv[64] := 0;
   tvv[65] := 0;
   tvv[66] := 0;
   tvv[67] := 0;
   tvv[68] := 0;
   tvv[69] := 0;
   tvv[70] := 0;
   tvv[71] := 0;
   tvv[72] := 0;
   tvv[73] := 0;
   tvv[74] := 0;
   tvv[75] := 0;
   tvv[76] := 0;
   tvv[77] := 0;
   tvv[78] := 0;
   tvv[79] := 0;
   tvv[80] := 0;
   tvv[81] := 0;
   tvv[82] := 0;
   tvv[83] := 0;
   tvv[84] := 0;
   tvv[85] := 0;
   tvv[86] := 0;
   tvv[87] := 0;
   tvv[88] := 0;
   tvv[89] := 0;
   tvv[90] := 0;
   tvv[91] := 0;
   tvv[92] := 0;
   tvv[93] := 0;
   tvv[94] := 0;
   tvv[95] := 0;
   tvv[96] := 0;
   tvv[97] := 0;
   tvv[98] := 0;
   tvv[99] := 0;
   spare[0] := 0;
   spare[1] := 0;
   spare[2] := 0;
   spare[3] := 0;
   spare[4] := 0;
   spare[5] := 0;
   spare[6] := 0;
   spare[7] := 0;
   spare[8] := 0;
   spare[9] := 0;
   spare[10] := 0;
   spare[11] := 0;
   spare[12] := 0;
   spare[13] := 0;
   spare[14] := 0;
   spare[15] := 0;
   spare[16] := 0;
   spare[17] := 0;
   spare[18] := 0;
   spare[19] := 0;
   spare[20] := 0;
   spare[21] := 0;
   spare[22] := 0;
   spare[23] := 0;
   spare[24] := 0;
   spare[25] := 0;
   spare[26] := 0;
   spare[27] := 0;
   spare[28] := 0;
   spare[29] := 0;
   spare[30] := 0;
   tach.ST := T#0MS;
   tach.PT := T#0MS;
   tach.RU := FALSE;
   tach.IN := FALSE;
   T_100ms.ST := T#-4D_23H_49M_55S_620MS;
   T_100ms.PT := T#100MS;
   T_100ms.RU := TRUE;
   T_100ms.IN := TRUE;
END_DATA_BLOCK

